// TIA Portal project "1905391_001_000" (V16) (continued)
FUNCTION_BLOCK "Material_Message"   // FB21, SCL
{ S7_Optimized_Access := 'TRUE' }
VERSION : 0.1
   VAR_INPUT
      adp_liberary : "ADP.Encoded.UDT";
   END_VAR
   VAR_IN_OUT
      hmi_interface : "HMI_Interface.UDT";
      led_interface : "LED_Interface.UDT";
   END_VAR
   VAR
      mode : String;
      old : Struct
         mode : String;
      END_STRUCT;
      set_mode : "Material_Message.Set_Mode";
      send_request : "Message.Request_Send";
      "Material_Message.Reset_Display_Driver" : "Material_Message.Reset_Display_Driver";
   END_VAR
BEGIN
   #set_mode(manual_request := #hmi_interface.connection_controls.material.send.operation_button_actuate,
             mode := #mode);

   IF #mode = "AUTOMATIC" THEN
       #"Material_Message.Reset_Display_Driver"(send_buffer := #led_interface.send_buffer,
                                                interface := #hmi_interface.materials);
       "Material_Message.Assemble_Automatic_Message"(adp_library := #adp_liberary,
                                                     interface := #hmi_interface.materials,
                                                     send_buffer := #led_interface.send_buffer);
   END_IF;

   IF #mode = "MANUAL" AND #mode <> #old.mode THEN
       "Material_Message.Assemble_Manual_Message"(adp_library := #adp_liberary,
                                                  send_buffer := #led_interface.send_buffer);
   END_IF;

   #old.mode := #mode;

   #send_request(manual_request := #hmi_interface.connection_controls.material.send.operation_button_actuate,
                 send_buffer := #led_interface.send_buffer,
                 send_request := #led_interface.requests.send);
END_FUNCTION_BLOCK

FUNCTION_BLOCK "Material_Message.Set_Mode"   // FB23, SCL
{ S7_Optimized_Access := 'TRUE' }
VERSION : 0.1
   VAR_INPUT
      manual_request : Bool;
      automatic_request : Bool;
   END_VAR
   VAR_IN_OUT
      mode : String;
   END_VAR
   VAR
      manual_delay : TOF_TIME;
      old : Struct
         in_manual_delay : Bool;
      END_STRUCT;
   END_VAR
   VAR_TEMP
      _in_manual_delay : Bool;
      _et : Time;
   END_VAR
   VAR CONSTANT
      DELAY : Time := T#15S;
   END_VAR
BEGIN
   #manual_delay(IN := #manual_request AND NOT #manual_delay.Q,
                 PT := #DELAY,
                 Q => #_in_manual_delay,
                 ET => #_et);

   IF NOT #_in_manual_delay THEN
       #mode := "AUTOMATIC";
       #old.in_manual_delay := #_in_manual_delay;
       RETURN;
   END_IF;

   #mode := "MANUAL";
   #old.in_manual_delay := #_in_manual_delay;
   RETURN;
END_FUNCTION_BLOCK

FUNCTION "Material_Message.Assemble_Automatic_Message" : Void   // FC166, SCL
{ S7_Optimized_Access := 'TRUE' }
VERSION : 0.1
   VAR_INPUT
      adp_library : "ADP.Encoded.UDT";
      interface : "Materials.HMI.UDT";
   END_VAR
   VAR_IN_OUT
      send_buffer : "ADP.Message_Buffer.UDT";
   END_VAR
   VAR_TEMP
      _count : UInt;
      _i : Int;
      _message : String;
      _rows : Array[0..8] of String;
      _send_buffer : "ADP.Message_Buffer.UDT";
   END_VAR
BEGIN
   REGION "MESSAGE HEADER"
       #_message := CONCAT_STRING(IN1 := #adp_library.file_system."00 Start of Header",
                                  IN2 := #adp_library.file_system."01 Address",
                                  IN3 := #adp_library.file_system."02 Start of Text",
                                  IN4 := #adp_library.file_system."03 Command & File",
                                  IN5 := #adp_library.formatting.size_and_face.normal_7);
   END_REGION


   REGION "TABLE ROWS"
       #_rows[0] := "Message.Assemble_Row"(adp_library := #adp_library,
                                           cell_0_value := 'HEAT',
                                           cell_0_color := #adp_library.formatting.color.yellow,
                                           cell_1_value := #interface.heat.cell_1_value,
                                           cell_1_color := '');

       #_rows[1] := "Message.Assemble_Row"(adp_library := #adp_library,
                                           cell_0_value := 'MATERIAL',
                                           cell_0_color := #adp_library.formatting.color.blue,
                                           cell_1_value := 'BAGS',
                                           cell_1_color := '');


       #_rows[2] := "Message.Assemble_Row"(adp_library := #adp_library,
                                           cell_0_value := 'MANGANESE',
                                           cell_0_color := #adp_library.formatting.color.white,
                                           cell_1_value := #interface.manganese.cell_1_value,
                                           cell_1_color := '');

       #_rows[3] := "Message.Assemble_Row"(adp_library := #adp_library,
                                           cell_0_value := 'SILICON',
                                           cell_0_color := '',
                                           cell_1_value := #interface.silicon.cell_1_value,
                                           cell_1_color := '');

       #_rows[4] := "Message.Assemble_Row"(adp_library := #adp_library,
                                           cell_0_value := 'CHROMIUM',
                                           cell_0_color := '',
                                           cell_1_value := #interface.chromium.cell_1_value,
                                           cell_1_color := '');

       #_rows[5] := "Message.Assemble_Row"(adp_library := #adp_library,
                                           cell_0_value := 'VANADIUM',
                                           cell_0_color := '',
                                           cell_1_value := #interface.vanadium.cell_1_value,
                                           cell_1_color := '');

       #_rows[6] := "Message.Assemble_Row"(adp_library := #adp_library,
                                           cell_0_value := 'NICKEL',
                                           cell_0_color := '',
                                           cell_1_value := #interface.nickel.cell_1_value,
                                           cell_1_color := '');

       #_rows[7] := "Message.Assemble_Row"(adp_library := #adp_library,
                                           cell_0_value := 'MOLYBDENUM',
                                           cell_0_color := '',
                                           cell_1_value := #interface.molybdenum.cell_1_value,
                                           cell_1_color := '');

       #_rows[8] := "Message.Assemble_Row"(adp_library := #adp_library,
                                           cell_0_value := #interface.custom.cell_0_value,
                                           cell_0_color := '',
                                           cell_1_value := #interface.custom.cell_1_value,
                                           cell_1_color := '');
       #_rows[8] := LEFT_STRING(IN := #_rows[8], L := LEN(#_rows[8]) - 1);
   END_REGION


   REGION "CONCAT HEADER AND ROWS"
       FOR #_i := 0 TO 8 DO
           #_message := CONCAT_STRING(IN1 := #_message, IN2 := #_rows[#_i]);
       END_FOR;
   END_REGION


   REGION "END OF MESSAGE"
       #_message := CONCAT_STRING(IN1 := #_message, IN2 := #adp_library.file_system."04 END");
   END_REGION


   REGION "RETURN"
       Strg_TO_Chars(Strg := #_message,
                     pChars := 0,
                     Cnt => #_count,
                     Chars := #send_buffer.me);
   END_REGION
END_FUNCTION

FUNCTION "Material_Message.Assemble_Manual_Message" : Void   // FC181, SCL
{ S7_Optimized_Access := 'TRUE' }
VERSION : 0.1
   VAR_INPUT
      adp_library : "ADP.Encoded.UDT";
   END_VAR
   VAR_IN_OUT
      send_buffer : "ADP.Message_Buffer.UDT";
   END_VAR
   VAR_TEMP
      _count : UInt;
      _i : Int;
      _message : String;
      _rows : Array[0..8] of String;
      _send_buffer : "ADP.Message_Buffer.UDT";
   END_VAR
BEGIN
   #_message := CONCAT_STRING(IN1 := #adp_library.file_system."00 Start of Header",
                              IN2 := #adp_library.file_system."01 Address",
                              IN3 := #adp_library.file_system."02 Start of Text",
                              IN4 := #adp_library.file_system."03 Command & File",
                              IN5 := 'MATERIAL COMMUNICATIONS TEST',
                              IN6 := #adp_library.file_system."04 END");


   Strg_TO_Chars(Strg := #_message,
                 pChars := 0,
                 Cnt => #_count,
                 Chars := #send_buffer.me);
END_FUNCTION

FUNCTION "Material_Message.Reset_Display" : Void   // FC194, SCL
{ S7_Optimized_Access := 'TRUE' }
VERSION : 0.1
   VAR_IN_OUT
      interface : "Materials.HMI.UDT";
   END_VAR
   VAR CONSTANT
      BLANK : String;
   END_VAR
BEGIN
   #interface.heat.cell_1_value := #BLANK;
   #interface.manganese.cell_1_value := #BLANK;
   #interface.silicon.cell_1_value := #BLANK;
   #interface.chromium.cell_1_value := #BLANK;
   #interface.vanadium.cell_1_value := #BLANK;
   #interface.nickel.cell_1_value := #BLANK;
   #interface.molybdenum.cell_1_value := #BLANK;
   #interface.custom.cell_1_value := #BLANK;
END_FUNCTION

// folder: material_sign

FUNCTION "Material_Sign.Set_Connection_Parameters" : Void   // FC123, SCL
{ S7_Optimized_Access := 'TRUE' }
VERSION : 0.1
   VAR_INPUT
      mode : String;
   END_VAR
   VAR_IN_OUT
      interface : "Connection_Parameters_HMI_Interface.UDT";
      saved : "Connection_Parameters.UDT";
   END_VAR
BEGIN
   IF #mode <> "MATERIAL" THEN
       RETURN;
   END_IF;
   "Connection_Parameters.Set_Parameters"(interface := #interface,
                                          saved :=#saved);
   RETURN;
END_FUNCTION

// folder: message

FUNCTION_BLOCK "Message.Detect_Change"   // FB22, SCL
{ S7_Optimized_Access := 'TRUE' }
VERSION : 0.1
   VAR_INPUT
      send_buffer : "ADP.Message_Buffer.UDT";
   END_VAR
   VAR_IN_OUT
      detected : Bool;
   END_VAR
   VAR
      old : Struct
         send_buffer : "ADP.Message_Buffer.UDT";
      END_STRUCT;
   END_VAR
BEGIN
   #detected := #send_buffer <> #old.send_buffer;
   #old.send_buffer := #send_buffer;
END_FUNCTION_BLOCK

FUNCTION_BLOCK "Message.Request_Send"   // FB24, SCL
{ S7_Optimized_Access := 'TRUE' }
VERSION : 0.1
   VAR_INPUT
      manual_request : Bool;
      send_buffer : "ADP.Message_Buffer.UDT";
   END_VAR
   VAR_IN_OUT
      send_request : Bool;
   END_VAR
   VAR
      "Message.Detect_Change" : "Message.Detect_Change";
   END_VAR
   VAR_TEMP
      _change_detected : Bool;
   END_VAR
BEGIN
   #"Message.Detect_Change"(send_buffer := #send_buffer,
                            detected := #_change_detected);
   IF #manual_request THEN
       #send_request := TRUE;
       RETURN;
   END_IF;
   IF #_change_detected THEN
       #send_request := TRUE;
       RETURN;
   END_IF;
   #send_request := FALSE;
   RETURN;
END_FUNCTION_BLOCK

FUNCTION "Message.Process_Color" : String   // FC11, SCL
{ S7_Optimized_Access := 'TRUE' }
VERSION : 0.1
   VAR_INPUT
      color : String;
   END_VAR
BEGIN
   IF LEN(#color) <> 0 THEN
       #"Message.Process_Color" := #color;
       RETURN;
   END_IF;
   #"Message.Process_Color" := '';
END_FUNCTION

FUNCTION "Message.Assemble_Row" : String   // FC167, SCL
{ S7_Optimized_Access := 'TRUE' }
VERSION : 0.1
   VAR_INPUT
      adp_library : "ADP.Encoded.UDT";
      cell_0_value : String;
      cell_0_color : String;
      cell_1_value : String;
      cell_1_color : String;
   END_VAR
   VAR_TEMP
      _cell_0 : String;
      _cell_0_color : String;
      _cell_1 : String;
      _cell_1_color : String;
      _return : String;
   END_VAR
BEGIN
   #_cell_0_color := "Message.Process_Color"(#cell_0_color);
   #_cell_0 := "String.Add_Leading"("Leading Character" := ' ',
                                    "Desired Length" := INT_TO_USINT(LEN(#cell_0_value)) + 1,
                                    "String" := #cell_0_value);
   #_cell_0 := "String.Add_Trailing"(value := #_cell_0,
                                     count := 12 - INT_TO_USINT(LEN(#_cell_0)),
                                     add_character := ' ');

   #_cell_1_color := "Message.Process_Color"(#cell_1_color);
   #_cell_1 := "String.Add_Leading"("Leading Character" := ' ',
                                    "Desired Length" := 7,
                                    "String" := #cell_1_value);
   #_cell_1 := "String.Add_Trailing"(value := #_cell_1,
                                     count := 1,
                                     add_character := ' ');

   #_return := CONCAT_STRING(IN1 := #_cell_0_color,
                             IN2 := #_cell_0,
                             IN3 := ' ',
                             IN4 := #_cell_1_color,
                             IN5 := #_cell_1,
                             IN6 := #adp_library.formatting.line_control.new_line);
   #"Message.Assemble_Row" := #_return;
END_FUNCTION

// folder: navigation

FUNCTION "Navigation.Initialize_Colors" : Void   // FC47, SCL
{ S7_Optimized_Access := 'TRUE' }
VERSION : 0.1
   VAR_IN_OUT
      navigation : "Navigation.HMI.UDT";
   END_VAR
BEGIN
   #navigation.background_animate := "Color.String_to_DInt"("BACKGROUND_COLOR");
   #navigation.bottom_line_animate := "Color.String_to_DInt"("DIVIDER_COLOR");
   #navigation.communications_status_animate := "Color.String_to_DInt"("OTHER_SCREEN_COLOR");
   #navigation.communications_status_cover_animate := "Color.String_to_DInt"("THIS_SCREEN_COLOR");
   #navigation.material_animate := "Color.String_to_DInt"("OTHER_SCREEN_COLOR");
   #navigation.material_cover_animate := "Color.String_to_DInt"("THIS_SCREEN_COLOR");
   #navigation.wire_animate := "Color.String_to_DInt"("THIS_SCREEN_COLOR");
   #navigation.wire_cover_animate := "Color.String_to_DInt"("THIS_SCREEN_COLOR");
END_FUNCTION

FUNCTION "Navigation.Wire_Animation" : Void   // FC48, SCL
{ S7_Optimized_Access := 'TRUE' }
VERSION : 0.1
   VAR_INPUT
      screen_number : Int;
   END_VAR
   VAR_IN_OUT
      navigation : "Navigation.HMI.UDT";
   END_VAR
   VAR_TEMP
      _color_off : DInt;
   END_VAR
BEGIN
   CASE #screen_number OF
       "WIRE_SCREEN_NUMBER":
           #_color_off := "Color.String_to_DInt"("THIS_SCREEN_COLOR");
       ELSE
           #_color_off := "Color.String_to_DInt"("OTHER_SCREEN_COLOR");
   END_CASE;
   "Bool.Animate"(signal := #navigation.wire_actuate,
                  color_on := "Color.String_to_DInt"("ACTUATE"),
                  color_off := #_color_off,
                  animation := #navigation.wire_animate);
END_FUNCTION

FUNCTION "Navigation.Initialize_Visibility" : Void   // FC60, SCL
{ S7_Optimized_Access := 'TRUE' }
VERSION : 0.1
   VAR_IN_OUT
      navigation : "Navigation.HMI.UDT";
   END_VAR
BEGIN
   #navigation.background_visible := TRUE;
   #navigation.bottom_line_visible := TRUE;
   #navigation.communications_status_cover_visible := FALSE;
   #navigation.communications_status_visible := TRUE;
   #navigation.material_cover_visible := FALSE;
   #navigation.material_visible := TRUE;
   #navigation.wire_cover_visible := TRUE;
   #navigation.wire_visible := TRUE;
END_FUNCTION

FUNCTION "Navigation.Initialize_Display" : Void   // FC61, SCL
{ S7_Optimized_Access := 'TRUE' }
VERSION : 0.1
   VAR_IN_OUT
      navigation : "Navigation.HMI.UDT";
   END_VAR
BEGIN
   "Navigation.Initialize_Colors"(#navigation);
   "Navigation.Initialize_Enable"(#navigation);
   "Navigation.Initialize_Visibility"(#navigation);
END_FUNCTION

FUNCTION "Navigation.Material_Animation" : Void   // FC66, SCL
{ S7_Optimized_Access := 'TRUE' }
VERSION : 0.1
   VAR_INPUT
      screen_number : Int;
   END_VAR
   VAR_IN_OUT
      navigation : "Navigation.HMI.UDT";
   END_VAR
   VAR_TEMP
      _color_off : DInt;
   END_VAR
BEGIN
   CASE #screen_number OF
       "MATERIAL_SCREEN_NUMBER":
           #_color_off := "Color.String_to_DInt"("THIS_SCREEN_COLOR");
       ELSE
           #_color_off := "Color.String_to_DInt"("OTHER_SCREEN_COLOR");
   END_CASE;
   "Bool.Animate"(signal := #navigation.material_actuate,
                  color_on := "Color.String_to_DInt"("ACTUATE"),
                  color_off := #_color_off,
                  animation := #navigation.material_animate);
END_FUNCTION

FUNCTION "Navigation.Initialize_Enable" : Void   // FC69, SCL
{ S7_Optimized_Access := 'TRUE' }
VERSION : 0.1
   VAR_IN_OUT
      navigation : "Navigation.HMI.UDT";
   END_VAR
BEGIN
   #navigation.communications_status_enable := TRUE;
   #navigation.material_enable := TRUE;
   #navigation.wire_enable := TRUE;
END_FUNCTION

FUNCTION "Navigation.Bottom_Cover_Animations" : Void   // FC73, SCL
{ S7_Optimized_Access := 'TRUE' }
VERSION : 0.1
   VAR_INPUT
      screen_number : Int;
   END_VAR
   VAR_IN_OUT
      navigation : "Navigation.HMI.UDT";
   END_VAR
BEGIN
   CASE #screen_number OF
       "MATERIAL_SCREEN_NUMBER":
           "Navigation.Connections_Screen_Hide_Bottom_Cover"(#navigation);
           "Navigation.Material_Screen_Show_Bottom_Cover"(#navigation);
           "Navigation.Wire_Screen_Hide_Bottom_Cover"(#navigation);
       "WIRE_SCREEN_NUMBER":
           "Navigation.Connections_Screen_Hide_Bottom_Cover"(#navigation);
           "Navigation.Material_Screen_Hide_Bottom_Cover"(#navigation);
           "Navigation.Wire_Screen_Show_Bottom_Cover"(#navigation);
       ELSE
           "Navigation.Connections_Screen_Show_Bottom_Cover"(#navigation);
           "Navigation.Material_Screen_Hide_Bottom_Cover"(#navigation);
           "Navigation.Wire_Screen_Hide_Bottom_Cover"(#navigation);
   END_CASE;
END_FUNCTION

FUNCTION "Navigation.Wire_Screen_Show_Bottom_Cover" : Void   // FC74, SCL
{ S7_Optimized_Access := 'TRUE' }
VERSION : 0.1
   VAR_IN_OUT
      navigation : "Navigation.HMI.UDT";
   END_VAR
BEGIN
   #navigation.wire_cover_visible := TRUE;
END_FUNCTION

FUNCTION "Navigation.Material_Screen_Show_Bottom_Cover" : Void   // FC75, SCL
{ S7_Optimized_Access := 'TRUE' }
VERSION : 0.1
   VAR_IN_OUT
      navigation : "Navigation.HMI.UDT";
   END_VAR
BEGIN
   #navigation.material_cover_visible := TRUE;
END_FUNCTION

FUNCTION "Navigation.Connections_Screen_Animation" : Void   // FC79, SCL
{ S7_Optimized_Access := 'TRUE' }
VERSION : 0.1
   VAR_INPUT
      screen_number : Int;
   END_VAR
   VAR_IN_OUT
      navigation : "Navigation.HMI.UDT";
   END_VAR
   VAR_TEMP
      _color_off : DInt;
   END_VAR
BEGIN
   CASE #screen_number OF
       "CONNECTION_CONTROLS_SCREEN_NUMBER":
           #_color_off := "Color.String_to_DInt"("THIS_SCREEN_COLOR");
       "CONNECTION_STATUS_DETAILS_SCREEN_NUMBER":
           #_color_off := "Color.String_to_DInt"("THIS_SCREEN_COLOR");
       "CONNECTION_PARAMETERS_SCREEN_NUMBER":
           #_color_off := "Color.String_to_DInt"("THIS_SCREEN_COLOR");
       ELSE
           #_color_off := "Color.String_to_DInt"("OTHER_SCREEN_COLOR");
   END_CASE;
   "Bool.Animate"(signal := #navigation.communications_status_actuate,
                  color_on := "Color.String_to_DInt"("ACTUATE"),
                  color_off := #_color_off,
                  animation := #navigation.communications_status_animate);
END_FUNCTION

FUNCTION "Navigation.Wire_Screen_Hide_Bottom_Cover" : Void   // FC80, SCL
{ S7_Optimized_Access := 'TRUE' }
VERSION : 0.1
   VAR_IN_OUT
      navigation : "Navigation.HMI.UDT";
   END_VAR
BEGIN
   #navigation.wire_cover_visible := FALSE;
END_FUNCTION

FUNCTION "Navigation.Connections_Screen_Show_Bottom_Cover" : Void   // FC81, SCL
{ S7_Optimized_Access := 'TRUE' }
VERSION : 0.1
   VAR_IN_OUT
      navigation : "Navigation.HMI.UDT";
   END_VAR
BEGIN
   #navigation.communications_status_cover_visible := TRUE;
END_FUNCTION

FUNCTION "Navigation.Connections_Screen_Hide_Bottom_Cover" : Void   // FC82, SCL
{ S7_Optimized_Access := 'TRUE' }
VERSION : 0.1
   VAR_IN_OUT
      navigation : "Navigation.HMI.UDT";
   END_VAR
BEGIN
   #navigation.communications_status_cover_visible := FALSE;
END_FUNCTION

FUNCTION "Navigation.Material_Screen_Hide_Bottom_Cover" : Void   // FC83, SCL
{ S7_Optimized_Access := 'TRUE' }
VERSION : 0.1
   VAR_IN_OUT
      navigation : "Navigation.HMI.UDT";
   END_VAR
BEGIN
   #navigation.material_cover_visible := FALSE;
END_FUNCTION

// folder: nibble

FUNCTION "Nibble.to_String" : String   // FC116, SCL
{ S7_Optimized_Access := 'TRUE' }
VERSION : 0.1
   VAR_INPUT
      value : Byte;
   END_VAR
   VAR_TEMP
      _nibble_as_int : Int;
      _ret : String;
   END_VAR
BEGIN
   #_nibble_as_int := BYTE_TO_INT(#value);
   CASE #_nibble_as_int OF
       0..9:
           #_ret := "String.Trim"("String.Strip_Sign"(INT_TO_STRING(#_nibble_as_int)));
       10:
           #_ret := 'A';
       11:
           #_ret := 'B';
       12:
           #_ret := 'C';
       13:
           #_ret := 'D';
       14:
           #_ret := 'E';
       15:
           #_ret := 'F';
   END_CASE;
   #"Nibble.to_String" := #_ret;
END_FUNCTION

// folder: row_custom

FUNCTION "Row_Custom.Animate_In_Focus" : Void   // FC9, SCL
{ S7_Optimized_Access := 'TRUE' }
VERSION : 0.1
   VAR_IN_OUT
      row_custom : "Row_Custom.UDT";
   END_VAR
BEGIN
   "Bool.Animate"(signal := #row_custom.cell_0_activate,
                  color_on := "Color.String_to_DInt"("SELECTED_INPUT_COLOR"),
                  color_off := "Color.String_to_DInt"("DESELECTED_INPUT_COLOR"),
                  animation := #row_custom.cell_0_animate);
   "Bool.Animate"(signal := #row_custom.cell_1_activate,
                  color_on := "Color.String_to_DInt"("SELECTED_INPUT_COLOR"),
                  color_off := "Color.String_to_DInt"("DESELECTED_INPUT_COLOR"),
                  animation := #row_custom.cell_1_animate);
END_FUNCTION

FUNCTION "Row_Custom.Hide" : Void   // FC41, SCL
{ S7_Optimized_Access := 'TRUE' }
VERSION : 0.1
   VAR_IN_OUT
      row_custom : "Row_Custom.UDT";
   END_VAR
   VAR CONSTANT
      MODE : Bool := FALSE;
   END_VAR
BEGIN
   #row_custom.background_visible := #MODE;
   #row_custom.cell_0_visible := #MODE;
   #row_custom.cell_1_visible := #MODE;
END_FUNCTION

FUNCTION "Row_Custom.Enable" : Void   // FC42, SCL
{ S7_Optimized_Access := 'TRUE' }
VERSION : 0.1
   VAR_IN_OUT
      row_custom : "Row_Custom.UDT";
   END_VAR
   VAR CONSTANT
      MODE : Bool := TRUE;
   END_VAR
BEGIN
   #row_custom.cell_0_enable := #MODE;
   #row_custom.cell_1_enable := #MODE;
END_FUNCTION

FUNCTION "Row_Custom.Initialize_Colors" : Void   // FC43, SCL
{ S7_Optimized_Access := 'TRUE' }
VERSION : 0.1
   VAR_IN_OUT
      row_custom : "Row_Custom.UDT";
   END_VAR
BEGIN
   #row_custom.background_animate := "Color.String_to_DInt"("BORDER_COLOR");
   #row_custom.cell_0_animate := "Color.String_to_DInt"("DESELECTED_INPUT_COLOR");
   #row_custom.cell_1_animate := "Color.String_to_DInt"("DESELECTED_INPUT_COLOR");
END_FUNCTION

FUNCTION "Row_Custom.Initialize" : Void   // FC44, SCL
{ S7_Optimized_Access := 'TRUE' }
VERSION : 0.1
   VAR_IN_OUT
      row_custom : "Row_Custom.UDT";
   END_VAR
BEGIN
   "Row_Custom.Show"(#row_custom);
   "Row_Custom.Enable"(#row_custom);
   "Row_Custom.Initialize_Colors"(#row_custom);
END_FUNCTION

FUNCTION "Row_Custom.Show" : Void   // FC64, SCL
{ S7_Optimized_Access := 'TRUE' }
VERSION : 0.1
   VAR_IN_OUT
      row_custom : "Row_Custom.UDT";
   END_VAR
   VAR CONSTANT
      MODE : Bool := TRUE;
   END_VAR
BEGIN
   #row_custom.background_visible := #MODE;
   #row_custom.cell_0_visible := #MODE;
   #row_custom.cell_1_visible := #MODE;
END_FUNCTION

FUNCTION "Row_Custom.Disable" : Void   // FC65, SCL
{ S7_Optimized_Access := 'TRUE' }
VERSION : 0.1
   VAR_IN_OUT
      row_custom : "Row_Custom.UDT";
   END_VAR
   VAR CONSTANT
      MODE : Bool := FALSE;
   END_VAR
BEGIN
   #row_custom.cell_0_enable := #MODE;
   #row_custom.cell_1_enable := #MODE;
END_FUNCTION

FUNCTION "Row_Custom.Reset_Input_Finished" : Void   // FC78, SCL
{ S7_Optimized_Access := 'TRUE' }
VERSION : 0.1
   VAR_IN_OUT
      input_finished : Bool;
   END_VAR
BEGIN
   #input_finished := FALSE;
END_FUNCTION

// folder: row_data

FUNCTION "Row_Data.Initialize_Colors" : Void   // FC1, SCL
{ S7_Optimized_Access := 'TRUE' }
VERSION : 0.1
   VAR_IN_OUT
      row_data : "Row_Data.UDT";
   END_VAR
BEGIN
   #row_data.background_animate := "Color.String_to_DInt"("BORDER_COLOR");
   #row_data.cell_0_animate := "Color.String_to_DInt"("LABEL_COLOR");
   #row_data.cell_1_animate := "Color.String_to_DInt"("DESELECTED_INPUT_COLOR");
END_FUNCTION

FUNCTION "Row_Data.Animate_In_Focus" : Void   // FC5, SCL
{ S7_Optimized_Access := 'TRUE' }
VERSION : 0.1
   VAR_IN_OUT
      row_data : "Row_Data.UDT";
   END_VAR
BEGIN
   "Bool.Animate"(signal := #row_data.cell_1_active,
                  color_on := "Color.String_to_DInt"("SELECTED_INPUT_COLOR"),
                  color_off := "Color.String_to_DInt"("DESELECTED_INPUT_COLOR"),
                  animation := #row_data.cell_1_animate);
END_FUNCTION

FUNCTION "Row_Data.Show" : Void   // FC6, SCL
{ S7_Optimized_Access := 'TRUE' }
VERSION : 0.1
   VAR_IN_OUT
      row_data : "Row_Data.UDT";
   END_VAR
   VAR CONSTANT
      MODE : Bool := TRUE;
   END_VAR
BEGIN
   #row_data.background_visible := #MODE;
   #row_data.cell_0_visible := #MODE;
   #row_data.cell_1_visible := #MODE;
END_FUNCTION

FUNCTION "Row_Data.Enable" : Void   // FC7, SCL
{ S7_Optimized_Access := 'TRUE' }
VERSION : 0.1
   VAR_IN_OUT
      row_data : "Row_Data.UDT";
   END_VAR
   VAR CONSTANT
      MODE : Bool := TRUE;
   END_VAR
BEGIN
   #row_data.cell_1_enable := #MODE;
END_FUNCTION

FUNCTION "Row_Data.Hide" : Void   // FC23, SCL
{ S7_Optimized_Access := 'TRUE' }
VERSION : 0.1
   VAR_IN_OUT
      row_data : "Row_Data.UDT";
   END_VAR
   VAR CONSTANT
      MODE : Bool := FALSE;
   END_VAR
BEGIN
   #row_data.background_visible := #MODE;
   #row_data.cell_0_visible := #MODE;
   #row_data.cell_1_visible := #MODE;
END_FUNCTION

FUNCTION "Row_Data.Disable" : Void   // FC24, SCL
{ S7_Optimized_Access := 'TRUE' }
VERSION : 0.1
   VAR_IN_OUT
      row_data : "Row_Data.UDT";
   END_VAR
   VAR CONSTANT
      MODE : Bool := FALSE;
   END_VAR
BEGIN
   #row_data.cell_1_enable := #MODE;
END_FUNCTION

FUNCTION "Row_Data.Initialize" : Void   // FC28, SCL
{ S7_Optimized_Access := 'TRUE' }
VERSION : 0.1
   VAR_IN_OUT
      row_data : "Row_Data.UDT";
   END_VAR
BEGIN
   "Row_Data.Enable"(#row_data);
   "Row_Data.Initialize_Colors"(#row_data);
   "Row_Data.Show"(#row_data);
END_FUNCTION

FUNCTION "Row_Data.Reset_Input_Finished" : Void   // FC77, SCL
{ S7_Optimized_Access := 'TRUE' }
VERSION : 0.1
   VAR_IN_OUT
      row_data : "Row_Data.UDT";
   END_VAR
BEGIN
   #row_data.cell_1_input_finished := FALSE;
END_FUNCTION

// folder: row_label

FUNCTION "Row_Label.Show" : Void   // FC38, SCL
{ S7_Optimized_Access := 'TRUE' }
VERSION : 0.1
   VAR_IN_OUT
      row_label : "Row_Label.UDT";
   END_VAR
   VAR CONSTANT
      MODE : Bool := TRUE;
   END_VAR
BEGIN
   #row_label.background_visible := #MODE;
   #row_label.cell_0_visible := #MODE;
   #row_label.cell_1_visible := #MODE;
END_FUNCTION

FUNCTION "Row_Label.Initialize" : Void   // FC39, SCL
{ S7_Optimized_Access := 'TRUE' }
VERSION : 0.1
   VAR_IN_OUT
      row_label : "Row_Label.UDT";
   END_VAR
BEGIN
   "Row_Label.Show"(#row_label);
   "Row_Label.Initialize_Colors"(#row_label);
END_FUNCTION

FUNCTION "Row_Label.Initialize_Colors" : Void   // FC40, SCL
{ S7_Optimized_Access := 'TRUE' }
VERSION : 0.1
   VAR_IN_OUT
      row_label : "Row_Label.UDT";
   END_VAR
BEGIN
   #row_label.background_animate := "Color.String_to_DInt"("BORDER_COLOR");
   #row_label.cell_0_animate := "Color.String_to_DInt"("LABEL_COLOR");
   #row_label.cell_1_animate := "Color.String_to_DInt"("LABEL_COLOR");
END_FUNCTION

FUNCTION "Row_Label.Hide" : Void   // FC63, SCL
{ S7_Optimized_Access := 'TRUE' }
VERSION : 0.1
   VAR_IN_OUT
      row_label : "Row_Label.UDT";
   END_VAR
   VAR CONSTANT
      MODE : Bool := FALSE;
   END_VAR
BEGIN
   #row_label.background_visible := #MODE;
   #row_label.cell_0_visible := #MODE;
   #row_label.cell_1_visible := #MODE;
END_FUNCTION

// folder: screen_background

FUNCTION "Screen_Background.Initialize" : Void   // FC70, SCL
{ S7_Optimized_Access := 'TRUE' }
VERSION : 0.1
   VAR_IN_OUT
      background : "Screen_Background.UDT";
   END_VAR
BEGIN
   "Screen_Background.Initialize_Color"(#background);
   "Screen_Background.Initialize_Visibility"(#background);
END_FUNCTION

FUNCTION "Screen_Background.Initialize_Color" : Void   // FC71, SCL
{ S7_Optimized_Access := 'TRUE' }
VERSION : 0.1
   VAR_IN_OUT
      background : "Screen_Background.UDT";
   END_VAR
BEGIN
   #background.color := "Color.String_to_DInt"("THIS_SCREEN_COLOR");
END_FUNCTION

FUNCTION "Screen_Background.Initialize_Visibility" : Void   // FC72, SCL
{ S7_Optimized_Access := 'TRUE' }
VERSION : 0.1
   VAR_IN_OUT
      background : "Screen_Background.UDT";
   END_VAR
BEGIN
   #background.visible := TRUE;
END_FUNCTION

// folder: sign

FUNCTION_BLOCK "Sign.Connection"   // FB16, SCL
{ S7_Optimized_Access := 'TRUE' }
VERSION : 0.1
   VAR_IN_OUT
      interface : "LED_Interface.UDT";
   END_VAR
   VAR
      manage_connection : "Connection.Manage_Connection";
   END_VAR
   VAR RETAIN
      tcon_param : TCON_Param;
   END_VAR
   VAR
      send : "Send";
   END_VAR
BEGIN
   #manage_connection(connection_parameters := #interface.connection_parameters,
                      requests := #interface.requests,
                      tcon_param := #tcon_param,
                      statuses := #interface.statuses);


   #send(send_buffer := #interface.send_buffer,
         requests := #interface.requests,
         tcon_param := #tcon_param,
         saved_status := #interface.statuses.send);
END_FUNCTION_BLOCK

// folder: string

FUNCTION "String.Drop_Last_Character" : String   // FC12, SCL
{ S7_Optimized_Access := 'TRUE' }
VERSION : 0.1
   VAR_INPUT
      value : String;
   END_VAR
BEGIN
   #"String.Drop_Last_Character" := LEFT_STRING(IN := #value,
                                                L := LEN(#value) - 1);
END_FUNCTION

FUNCTION "String.Find" : Int   // FC18, SCL
{ S7_Optimized_Access := 'TRUE' }
VERSION : 0.1
   VAR_INPUT
      search_for : String;
      search_in : String;
   END_VAR
BEGIN
   #"String.Find" := FIND(IN1 := #search_in, IN2 := #search_for);
END_FUNCTION

FUNCTION "String.Strip_Sign" : String   // FC20, SCL
{ S7_Optimized_Access := 'TRUE' }
VERSION : 0.1
   VAR_INPUT
      "string" : String;
   END_VAR
   VAR_TEMP
      Length : Int;
      "String Box" : String;
      "Test Character" : String;
   END_VAR
   VAR CONSTANT
      "+" : Char := '+';
      "-" : Char := '-';
   END_VAR
BEGIN
   #"String Box" := #string;
   #"Test Character" := LEFT_STRING(IN := #"String Box",
                                    L := 1);
   IF #"Test Character" = #"+" OR #"Test Character" = #"-" THEN
       #Length := LEN(#"String Box");
       #"String Box" := RIGHT_STRING(IN := #"String Box", L := #Length - 1);

   END_IF;
   #"String.Strip_Sign" := #"String Box";
END_FUNCTION

FUNCTION "String.Trim" : String   // FC21, SCL
{ S7_Optimized_Access := 'TRUE' }
AUTHOR : Machado
FAMILY : String
VERSION : 1.0
// removes leading and trailing whitespace from input string
   VAR_INPUT
      "string" : String;
   END_VAR
   VAR_TEMP
      ret : String;
   END_VAR
   VAR CONSTANT
      space : String := ' ';
   END_VAR
BEGIN
   #ret := #string;
   WHILE LEFT(IN := #ret, L := 1) = #space DO
       #ret := RIGHT(IN := #ret, L := LEN(#ret) - 1);
   END_WHILE;
   WHILE RIGHT(IN := #ret, L := 1) = #space DO
       #ret := LEFT(IN := #ret, L := LEN(#ret) - 1);
   END_WHILE;
   #"String.Trim" := #ret;
END_FUNCTION

FUNCTION "String.Upper" : String   // FC22, SCL
{ S7_Optimized_Access := 'TRUE' }
AUTHOR : Machado
FAMILY : String
VERSION : 1.0
// returns the input string converted to all upper case
   VAR_INPUT
      "string" : String;
   END_VAR
   VAR_TEMP
      "type" : Bool;
      stringBox : String;
      status : Int;
      charArr : Array[0..255] of Char;
      cntChar : UInt;
      pChar : Int;
   END_VAR
   VAR CONSTANT
      asciiLow : Char := 'a';
      asciiHigh : Char := 'z';
      asciiCaseOffset : Int := 32;
   END_VAR
BEGIN
   Strg_TO_Chars(Strg := #string,
                 pChars := 0,
                 Cnt => #cntChar,
                 Chars := #charArr);

   FOR #pChar := 0 TO UINT_TO_INT(#cntChar) - 1 DO
       IF #asciiLow <= #charArr[#pChar] AND #charArr[#pChar] <= #asciiHigh THEN
           #charArr[#pChar] := INT_TO_CHAR(CHAR_TO_INT(#charArr[#pChar]) - #asciiCaseOffset);
       END_IF;
   END_FOR;

   Chars_TO_Strg(Chars := #charArr,
                 pChars := 0,
                 Cnt := #cntChar,
                 Strg => #stringBox);

   #"String.Upper" := #stringBox;
END_FUNCTION

FUNCTION "String.Split_Multiple" : Void   // FC26, SCL
{ S7_Optimized_Access := 'TRUE' }
VERSION : 0.1
   VAR_INPUT
      string_in : String;
      delimeters : Array[*] of String;
      pointer : Int;
   END_VAR
   VAR_OUTPUT
      substrings : Array[*] of String;
   END_VAR
   VAR_TEMP
      _i : Int;
      _position : Int;
      _return : String;
      _split : String;
   END_VAR
BEGIN
   REGION "GET POSITION OF DELIMETER IN STRING"
       #_position := "String.Find_Multiple.Breadth"(body := #string_in,
                                                    terms := #delimeters);
   END_REGION

   REGION "BASE CASE"
       IF #_position = 0 THEN
           #substrings[#pointer] := #string_in;
           "String.Split_Multiple.Clean_Output"("pointer" := #pointer + 1,
                                                substrings := #substrings);
           RETURN;
       END_IF;
   END_REGION


   REGION "RECURSIVE CASE"
       #substrings[#pointer] := LEFT(IN := #string_in, L := #_position);
       "String.Split_Multiple"(string_in := RIGHT(IN := #string_in, L := LEN(#string_in) - #_position),
                               delimeters := #delimeters,
                               "pointer" := #pointer + 1,
                               substrings => #substrings);
   END_REGION
END_FUNCTION

FUNCTION "String.Split_Single" : Void   // FC33, SCL
{ S7_Optimized_Access := 'TRUE' }
VERSION : 0.1
   VAR_INPUT
      string_in : String;
      delimeter : String;
      pointer : Int;
   END_VAR
   VAR_IN_OUT
      sub_strings : Array[*] of String;
   END_VAR
   VAR_TEMP
      _split : String;
      _position : Int;
      _return : String;
   END_VAR
BEGIN
   REGION "GET POSITION OF DELIMETER IN STRING"
       #_position := FIND(IN1 := #string_in,
                          IN2 := #delimeter);
   END_REGION

   REGION "BASE CASE"
       IF #_position = 0 THEN
           #sub_strings[#pointer] := #string_in;
           RETURN;
       END_IF;
   END_REGION


   REGION "RECURSIVE CASE"
       #sub_strings[#pointer] := LEFT(IN := #string_in, L := #_position - 1);
       "String.Split_Single"(string_in := RIGHT(IN := #string_in, L := LEN(#string_in) - #_position),
                             delimeter := #delimeter,
                             "pointer" := #pointer + 1,
                             sub_strings := #sub_strings);
   END_REGION
END_FUNCTION

FUNCTION "String.Find_Multiple.Breadth" : Int   // FC34, SCL
{ S7_Optimized_Access := 'TRUE' }
VERSION : 0.1
   VAR_INPUT
      body : String;
      terms : Array[*] of String;
   END_VAR
   VAR_TEMP
      _i : Int;
      _length : UDInt;
      _min : Int;
      _position : Int;
   END_VAR
   VAR CONSTANT
      BLANK : String;
   END_VAR
BEGIN
   (* 
       Depth first search of 'body' for first occurance of any element of 'terms'.
       For depth first search use WString.Find_Multiple.Depth.
       Returns character postion in the string (1 indexed).
       E.G.: 
           - body := WSTRING#'today?'
           - terms := <WSTRING#>['?', 'ay']
           - returns --> 6
       E.G.:
           - body := WSTRING#'today?'
           - terms := <WSTRING#>['ay', '?']
           - returns --> 4
   *)

   #_length := "Any.Array.Length"(#terms);

   IF #_length = 0 OR #body = #BLANK THEN
       #"String.Find_Multiple.Breadth" := 0;
       RETURN;
   END_IF;

   FOR #_i := 0 TO UDINT_TO_INT(#_length) - 1 DO
       #_position := FIND(IN1 := #body,
                          IN2 := #terms[#_i]);
       IF #_position = 0 THEN
           CONTINUE;
       END_IF;
       IF #_position < #_min OR #_min = 0 THEN
           #_min := #_position;
       END_IF;
   END_FOR;

   #"String.Find_Multiple.Breadth" := #_min;
END_FUNCTION

FUNCTION "String.Split_Multiple.Clean_Output" : Void   // FC35, SCL
{ S7_Optimized_Access := 'TRUE' }
VERSION : 0.1
   VAR_INPUT
      pointer : Int;
   END_VAR
   VAR_IN_OUT
      substrings : Array[*] of String;
   END_VAR
   VAR_TEMP
      _i : Int;
   END_VAR
   VAR CONSTANT
      BLANK : String;
   END_VAR
BEGIN
   FOR #_i := #"pointer" TO UDINT_TO_INT("Any.Array.Length"(#substrings)) - 1 DO
       #substrings[#_i] := #BLANK;
   END_FOR;
END_FUNCTION

FUNCTION "String.Search_Array" : Int   // FC50, SCL
{ S7_Optimized_Access := 'TRUE' }
VERSION : 0.1
   VAR_INPUT
      "array" : Array[*] of String;
      search_term : String;
   END_VAR
   VAR_TEMP
      _i : Int;
      _length : Int;
   END_VAR
BEGIN
   REGION "SEARCH ARRAY"    
       #_length := UDINT_TO_INT("Any.Array.Length"(#array)) - 1;
       FOR #_i := 0 TO #_length DO
           IF #array[#_i] = #search_term THEN
               #"String.Search_Array" := #_i;
               RETURN;
           END_IF;
       END_FOR;
   END_REGION

   REGION "RETURN"
       #"String.Search_Array" := "NULL_TOKEN";
       RETURN;
   END_REGION
END_FUNCTION

FUNCTION "String.Reverse_Array" : Void   // FC51, SCL
{ S7_Optimized_Access := 'TRUE' }
VERSION : 0.1
   VAR_INPUT
      null_token : String;
   END_VAR
   VAR_IN_OUT
      string_array : Array[*] of String;
   END_VAR
   VAR_TEMP
      _has_data_count : Int;
      _i : Int;
      _p_swap : Int;
      _temp : String;
   END_VAR
   VAR CONSTANT
      NOT_FOUND : Int := -1;
   END_VAR
BEGIN
   REGION "CHECK FOR FIRST EMPTY POSITION"
       #_has_data_count := "String.Search_Array"(array := #string_array,
                                                 search_term := #null_token);
   END_REGION


   REGION "EXIT ON EMPTY ARRAY"
       IF #_has_data_count = 0 THEN
           RETURN;
       END_IF;
   END_REGION


   REGION "ARRAY IS FULL"
       IF #_has_data_count = #NOT_FOUND THEN
           #_has_data_count := UDINT_TO_INT("Any.Array.Length"(#string_array));
       END_IF;
   END_REGION


   REGION "ADJUST TO ZERO INDEX"
       #_has_data_count -= 1;
   END_REGION


   REGION "SWAP ELEMENTS"
       FOR #_i := 0 TO #_has_data_count / 2 DO
           #_p_swap := #_has_data_count - #_i;
           #_temp := #string_array[#_i];
           #string_array[#_i] := #string_array[#_p_swap];
           #string_array[#_p_swap] := #_temp;
       END_FOR;
   END_REGION


   REGION "DONE"
       RETURN;
   END_REGION
END_FUNCTION

FUNCTION "String.Is_Numeric" : Bool   // FC58, SCL
{ S7_Optimized_Access := 'TRUE' }
VERSION : 0.1
   VAR_INPUT
      "string" : String;
   END_VAR
   VAR_TEMP
      _string : String;
   END_VAR
BEGIN
   #_string := #string;
   WHILE LEN(#_string) > 0 DO
       IF NOT "Char.Is_Numeric"(STRING_TO_CHAR(LEFT_STRING(IN := #_string, L := 1))) THEN
           #"String.Is_Numeric" := FALSE;
           RETURN;
       END_IF;
       #_string := "String.Slice_Right"("string" := #_string,
                                        start_at := 1);
   END_WHILE;
   #"String.Is_Numeric" := TRUE;
   RETURN;
END_FUNCTION

FUNCTION "String.Slice_Right" : String   // FC59, SCL
{ S7_Optimized_Access := 'TRUE' }
VERSION : 0.1
   VAR_INPUT
      "string" : String;
      start_at : Int;
   END_VAR
   VAR_TEMP
      _length : Int;
   END_VAR
BEGIN
   #"String.Slice_Right" := RIGHT_STRING(IN := #string,
                                         L := LEN(#string) - #start_at);
END_FUNCTION

FUNCTION "String.Count" : Int   // FC62, SCL
{ S7_Optimized_Access := 'TRUE' }
VERSION : 0.1
   VAR_INPUT
      space : String;   // count term ocuurances in space
      term : String;
   END_VAR
   VAR_TEMP
      _count : Int;
      _position : Int;
      _space : String;
   END_VAR
BEGIN
   #_space := #space;
   #_position := FIND(IN1 := #_space,
                      IN2 := #term);
   IF #_position = 0 THEN
       #"String.Count" := 0;
       RETURN;
   END_IF;
   WHILE #_position > 0 DO
       #_count += 1;
       #_space := RIGHT(IN := #_space,
                        L := LEN(#_space) - #_position);
       #_position := FIND(IN1 := #_space,
                          IN2 := #term);
   END_WHILE;
   #"String.Count" := #_count;
   RETURN;
END_FUNCTION

FUNCTION "String.Center_Pad_Right" : String   // FC99, SCL
{ S7_Optimized_Access := 'TRUE' }
VERSION : 0.1
   VAR_INPUT
      value : String;
      spaces : USInt;
   END_VAR
   VAR_TEMP
      _length : USInt;
      _left : USInt;
      _right : USInt;
      _return : String;
   END_VAR
BEGIN
   #_length := INT_TO_USINT(LEN(#value));
   IF #_length > #spaces THEN
       #"String.Center_Pad_Right" := #value;
   END_IF;
   #_left := (#spaces - #_length) / 2;
   #_right := #_left;
   IF (#spaces - #_length) MOD 2 <> 0 THEN
       #_right += 1;
   END_IF;
   #_return := "String.Add_Leading"("Leading Character" := ' ',
                                    "Desired Length" := #_length + #_left,
                                    "String" := #value);
   #_return := "String.Add_Trailing"(value := #_return,
                                     count := #_right,
                                     add_character := ' ');
   #"String.Center_Pad_Right" := #_return;
END_FUNCTION

FUNCTION "String.Add_Leading" : String   // FC100, SCL
{ S7_Optimized_Access := 'TRUE' }
VERSION : 0.1
   VAR_INPUT
      "Leading Character" : Char;
      "Desired Length" : USInt;
      "String" : String;
   END_VAR
   VAR_TEMP
      Length : Int;
      "String Box" : String;
   END_VAR
BEGIN
   #"String Box" := #String;
   #Length := LEN(#"String Box");

   WHILE #Length < #"Desired Length" DO
       #"String Box" := CONCAT_STRING(IN1 := #"Leading Character",
                                      IN2 := #"String Box");
       #Length := LEN(#"String Box");
   END_WHILE;

   #"String.Add_Leading" := #"String Box";
END_FUNCTION

FUNCTION "String.Add_Trailing" : String   // FC101, SCL
{ S7_Optimized_Access := 'TRUE' }
VERSION : 0.1
   VAR_INPUT
      value : String;
      count : Int;
      add_character : Char;
   END_VAR
   VAR_TEMP
      _i : Int;
      _return : String;
   END_VAR
BEGIN
   IF #count <= 0 THEN
       #"String.Add_Trailing" := #value;
   END_IF;
   #_return := #value;
   FOR #_i := 0 TO #count - 1 DO
       #_return := CONCAT_STRING(IN1 := #_return, IN2 := CHAR_TO_STRING(#add_character));
   END_FOR;
   #"String.Add_Trailing" := #_return;
END_FUNCTION

FUNCTION "String.to_REM_STADDR" : Void   // FC102, SCL
{ S7_Optimized_Access := 'TRUE' }
VERSION : 0.1
   VAR_INPUT
      ip_address : String;   // use '.' or '_' to delimit octets
   END_VAR
   VAR_IN_OUT
      REM_STADDR : Array[1..6] of USInt;
   END_VAR
   VAR_TEMP
      _delimeters : Array[0..1] of String;
      _i : Int;
      _substrings : Array[0..3] of String;
   END_VAR
BEGIN
   #_delimeters[0] := '.';
   #_delimeters[1] := '_';
   "String.Split_Multiple"(string_in := #ip_address,
                           delimeters := #_delimeters,
                           "pointer" := 0,
                           substrings => #_substrings);
   FOR #_i := 1 TO 4 DO
       #REM_STADDR[#_i] := STRING_TO_USINT(#_substrings[#_i - 1]);
   END_FOR;
END_FUNCTION

FUNCTION "String.to_REM_TSAP_ID" : Void   // FC103, SCL
{ S7_Optimized_Access := 'TRUE' }
VERSION : 0.1
   VAR_INPUT
      port_number : String;
   END_VAR
   VAR_IN_OUT
      REM_TSAP_ID : Array[1..16] of Byte;
   END_VAR
   VAR_TEMP
      _as_uint : UInt;
   END_VAR
BEGIN
   #_as_uint := STRING_TO_UINT(#port_number);
   #REM_TSAP_ID[1] := #_as_uint.%B1;
   #REM_TSAP_ID[2] := #_as_uint.%B0;
END_FUNCTION

FUNCTION "String.Center_Pad_Left" : String   // FC182, SCL
{ S7_Optimized_Access := 'TRUE' }
VERSION : 0.1
   VAR_INPUT
      value : String;
      spaces : USInt;
   END_VAR
   VAR_TEMP
      _length : USInt;
      _left : USInt;
      _right : USInt;
      _return : String;
   END_VAR
BEGIN
   #_length := INT_TO_USINT(LEN(#value));
   IF #_length > #spaces THEN
       #"String.Center_Pad_Left" := #value;
   END_IF;
   #_left := (#spaces - #_length) / 2;
   #_right := #_left;
   IF (#spaces - #_length) MOD 2 <> 0 THEN
       #_left += 1;
   END_IF;
   #_return := "String.Add_Leading"("Leading Character" := ' ',
                                    "Desired Length" := #_length + #_left,
                                    "String" := #value);
   #_return := "String.Add_Trailing"(value := #_return,
                                     count := #_right,
                                     add_character := ' ');
   #"String.Center_Pad_Left" := #_return;
END_FUNCTION

FUNCTION "String.Array.Is_Element" : Bool   // FC195, SCL
{ S7_Optimized_Access := 'TRUE' }
VERSION : 0.1
   VAR_INPUT
      search_term : String;
      search_array : Array[*] of String;
   END_VAR
   VAR_TEMP
      _i : Int;
      _length_search_array : UDInt;
   END_VAR
BEGIN
   #_length_search_array := "Any.Array.Length"(#search_array);
   FOR #_i := 0 TO UDINT_TO_INT(#_length_search_array - 1) DO
       IF #search_term = #search_array[#_i] THEN
           #"String.Array.Is_Element" := TRUE;
           RETURN;
       END_IF;
   END_FOR;
   #"String.Array.Is_Element" := FALSE;
END_FUNCTION

FUNCTION "String.Word_Wrap" : String   // FC197, SCL
{ S7_Optimized_Access := 'TRUE' }
VERSION : 0.1
   VAR_INPUT
      delimeters : Array[*] of String;
      line_length : Int;
      value : String;
   END_VAR
   VAR_TEMP
      _i : Int;
      _substring_length : Int;
      _wstring_in_length : Int;
      _pointer_substrings : Int;
      _substring : String;
      _position_of_last_delimeter : Int;
      _recurse : Bool;
      _string_split_right : String;
   END_VAR
   VAR CONSTANT
      BLANK : String;
      NEW_LINE : String := '$L';
   END_VAR
BEGIN
   #_wstring_in_length := LEN(#value);

   IF #line_length = 0 THEN
       #"String.Word_Wrap" := #BLANK;
       RETURN;
   END_IF;

   FOR #_i := 1 TO #_wstring_in_length DO

       #_substring := CONCAT_STRING(IN1 := #_substring,
                                     IN2 := #value[#_i]);
       #_substring_length := LEN(#_substring);

       IF "String.Array.Is_Element"(search_term := #value[#_i], search_array := #delimeters) THEN
           #_position_of_last_delimeter := #_i;
       END_IF;

       IF #value[#_i] = #NEW_LINE THEN
           #_substring := LEFT_STRING(IN := #_substring,
                                       L := #_substring_length - 1);
           #_string_split_right := RIGHT_STRING(IN := #value,
                                                 L := #_wstring_in_length - #_i);
           #_recurse := TRUE;
       END_IF;

       IF (#_substring_length = #line_length) AND (#_position_of_last_delimeter <> 0) THEN
           #_substring := LEFT_STRING(IN := #_substring,
                                       L := #_position_of_last_delimeter);
           #_string_split_right := RIGHT_STRING(IN := #value,
                                                 L := #_wstring_in_length - #_position_of_last_delimeter);
           #_recurse := TRUE;
       END_IF;

       IF (#_substring_length = #line_length) AND (#_position_of_last_delimeter = 0) THEN
           #_string_split_right := RIGHT_STRING(IN := #value,
                                                 L := #_wstring_in_length - #_substring_length);
           #_recurse := TRUE;
       END_IF;

       IF #_recurse THEN
           #_substring := CONCAT_STRING(IN1 := "String.Trim"(#_substring),
                                         IN2 := #NEW_LINE,
                                         IN3 := "String.Word_Wrap"(delimeters := #delimeters,
                                                                    line_length := #line_length,
                                                                    value := #_string_split_right));
           #"String.Word_Wrap" := #_substring;
           RETURN;
       END_IF;

   END_FOR;

   #"String.Word_Wrap" := "String.Trim"(#_substring);
END_FUNCTION

// folder: tcpip_connection

FUNCTION_BLOCK "Connection.Manage_Connection"   // FB10, SCL
{ S7_Optimized_Access := 'TRUE' }
VERSION : 0.1
   VAR_INPUT
      connection_parameters : "Connection_Parameters.UDT";
   END_VAR
   VAR_IN_OUT
      requests : "Connection_Requests.UDT";
      tcon_param : TCON_Param;
      statuses : "Connection_Statuses.UDT";
   END_VAR
   VAR
      connect : "Connect";
      disconnect : "Disconnect";
      old : Struct
         connection_parameters : "Connection_Parameters.UDT";
      END_STRUCT;
      reset : "Reset";
      diagnostics : "Diagnostics";
   END_VAR
BEGIN
   IF "FirstScan" THEN
       "Connection.Load_TCON_Param"(interface := #connection_parameters,
                                    tcon_param := #tcon_param);
   END_IF;


   IF #connection_parameters <> #old.connection_parameters THEN
       "Connection.Load_TCON_Param"(interface := #connection_parameters,
                                    tcon_param := #tcon_param);
   END_IF;
   #old.connection_parameters := #connection_parameters;

   #connect(tcon_param := #tcon_param,
            requests := #requests,
            saved_status := #statuses.connect);


   #disconnect(tcon_param := #tcon_param,
               requests := #requests,
               saved_status := #statuses.disconnect);


   #reset(tcon_param := #tcon_param,
          requests := #requests);


   #diagnostics(tcon_param := #tcon_param,
                requests := #requests);
END_FUNCTION_BLOCK

FUNCTION "Connection.Initialize_Parameters" : Void   // FC104, SCL
{ S7_Optimized_Access := 'TRUE' }
VERSION : 0.1
   VAR_INPUT
      interface : "Connection_Parameters.UDT";
   END_VAR
   VAR_IN_OUT
      tcon_param : TCON_Param;
   END_VAR
BEGIN
   IF "FirstScan" THEN
       "Connection.Load_TCON_Param"(interface := #interface,
                                    tcon_param := #tcon_param);

   END_IF;
END_FUNCTION

FUNCTION "Connection.Load_TCON_Param" : Void   // FC137, SCL
{ S7_Optimized_Access := 'TRUE' }
VERSION : 0.1
   VAR_INPUT
      interface : "Connection_Parameters.UDT";
   END_VAR
   VAR_IN_OUT
      tcon_param : TCON_Param;
   END_VAR
BEGIN
   #tcon_param.ID := #interface.id;
   "String.to_REM_STADDR"(ip_address := #interface.ip_address,
                          REM_STADDR := #tcon_param.REM_STADDR);
   "String.to_REM_TSAP_ID"(port_number := #interface.port_number,
                           REM_TSAP_ID := #tcon_param.REM_TSAP_ID);
END_FUNCTION

// folder: tcpip_connection/connect

